REGION Network 15 (SCL): Calculate alarm statuses
   #ST_xStoppingFaults :=  #tALM.tS.xAxisNotAvail OR 
                               #tALM.tS.xInpInstallation OR 
                               #tALM.tS.xAuxPower OR 
                               #tALM.tS.xAreaSafety OR 
                               #tALM.tS.xOverstroke OR 
                               #tALM.tS.xExternInputPower OR 
                               #tALM.tS.xCarriageCutOut OR 
                               #tALM.tS.xDriveTrip OR 
                               #tALM.tS.xDriveNotEnabled OR 
                               #tALM.tS.xAxisNotReady OR 
                               #tALM.tS.xDriveNotReady OR 
                               #tALM.tS.xAxisNotSyncro OR 
                               #tALM.tS.xSpare_12 OR 
                               #tALM.tS.xSpare_13 OR 
                               #tALM.tS.xSpare_14 OR 
                               #tALM.tS.xSpare_15 OR 
                               #tALM.tS.xSpare_16 OR 
                               #tALM.tS.xSpare_17 OR 
                               #tALM.tS.xSpare_18 OR 
                               #tALM.tS.xSpare_19 OR 
                               #tALM.tS.xSpare_20 OR 
                               #tALM.tS.xSpare_21 OR 
                               #tALM.tS.xSpare_22 OR 
                               #tALM.tS.xSpare_23 OR 
                               #tALM.tS.xSpare_24 OR 
                               #tALM.tS.xSpare_25 OR 
                               #tALM.tS.xSpare_26 OR 
                               #tALM.tS.xSpare_27 OR 
                               #tALM.tS.xSpare_28 OR 
                               #tALM.tS.xSpare_29 OR 
                               #tALM.tS.xSpare_30 OR 
                               #tALM.tS.xSpare_31;

   #ST_xFaults := #tALM.tF.xSpare_0 OR
   #tALM.tF.xSpare_1 OR
   #tALM.tF.xSpare_2 OR
   #tALM.tF.xSpare_3 OR
   #tALM.tF.xSpare_4 OR
   #tALM.tF.xSpare_5 OR
   #tALM.tF.xSpare_6 OR
   #tALM.tF.xSpare_7 OR
   #tALM.tF.xSpare_8 OR
   #tALM.tF.xSpare_9 OR
   #tALM.tF.xSpare_10 OR
   #tALM.tF.xSpare_11 OR
   #tALM.tS.xSpare_12 OR
   #tALM.tS.xSpare_13 OR
   #tALM.tS.xSpare_14 OR
   #tALM.tS.xSpare_15 OR
   #tALM.tS.xSpare_16 OR
   #tALM.tS.xSpare_17 OR
   #tALM.tS.xSpare_18 OR
   #tALM.tS.xSpare_19 OR
   #tALM.tS.xSpare_20 OR
   #tALM.tS.xSpare_21 OR
   #tALM.tS.xSpare_22 OR
   #tALM.tS.xSpare_23 OR
   #tALM.tS.xSpare_24 OR
   #tALM.tS.xSpare_25 OR
   #tALM.tS.xSpare_26 OR
   #tALM.tS.xSpare_27 OR
   #tALM.tS.xSpare_28 OR
   #tALM.tS.xSpare_29 OR
   #tALM.tS.xSpare_30 OR
   #tALM.tS.xSpare_31;

   #ST_xWarnings := #tALM.tW.xSpare_0 OR
   #tALM.tW.xSpare_1 OR
   #tALM.tW.xSpare_2 OR
   #tALM.tW.xSpare_3 OR
   #tALM.tW.xSpare_4 OR
   #tALM.tW.xSpare_5 OR
   #tALM.tW.xSpare_6 OR
   #tALM.tW.xSpare_7 OR
   #tALM.tW.xSpare_8 OR
   #tALM.tW.xSpare_9 OR
   #tALM.tW.xSpare_10 OR
   #tALM.tW.xSpare_11 OR
   #tALM.tW.xSpare_12 OR
   #tALM.tW.xSpare_13 OR
   #tALM.tW.xSpare_14 OR
   #tALM.tW.xSpare_15 OR
   #tALM.tW.xSpare_16 OR
   #tALM.tW.xSpare_17 OR
   #tALM.tW.xSpare_18 OR
   #tALM.tW.xSpare_19 OR
   #tALM.tW.xSpare_20 OR
   #tALM.tW.xSpare_21 OR
   #tALM.tW.xSpare_22 OR
   #tALM.tW.xSpare_23 OR
   #tALM.tW.xSpare_24 OR
   #tALM.tW.xSpare_25 OR
   #tALM.tW.xSpare_26 OR
   #tALM.tW.xSpare_27 OR
   #tALM.tW.xSpare_28 OR
   #tALM.tW.xSpare_29 OR
   #tALM.tW.xSpare_30 OR
   #tALM.tW.xSpare_31;
END_REGION

REGION Network 16: Output enable
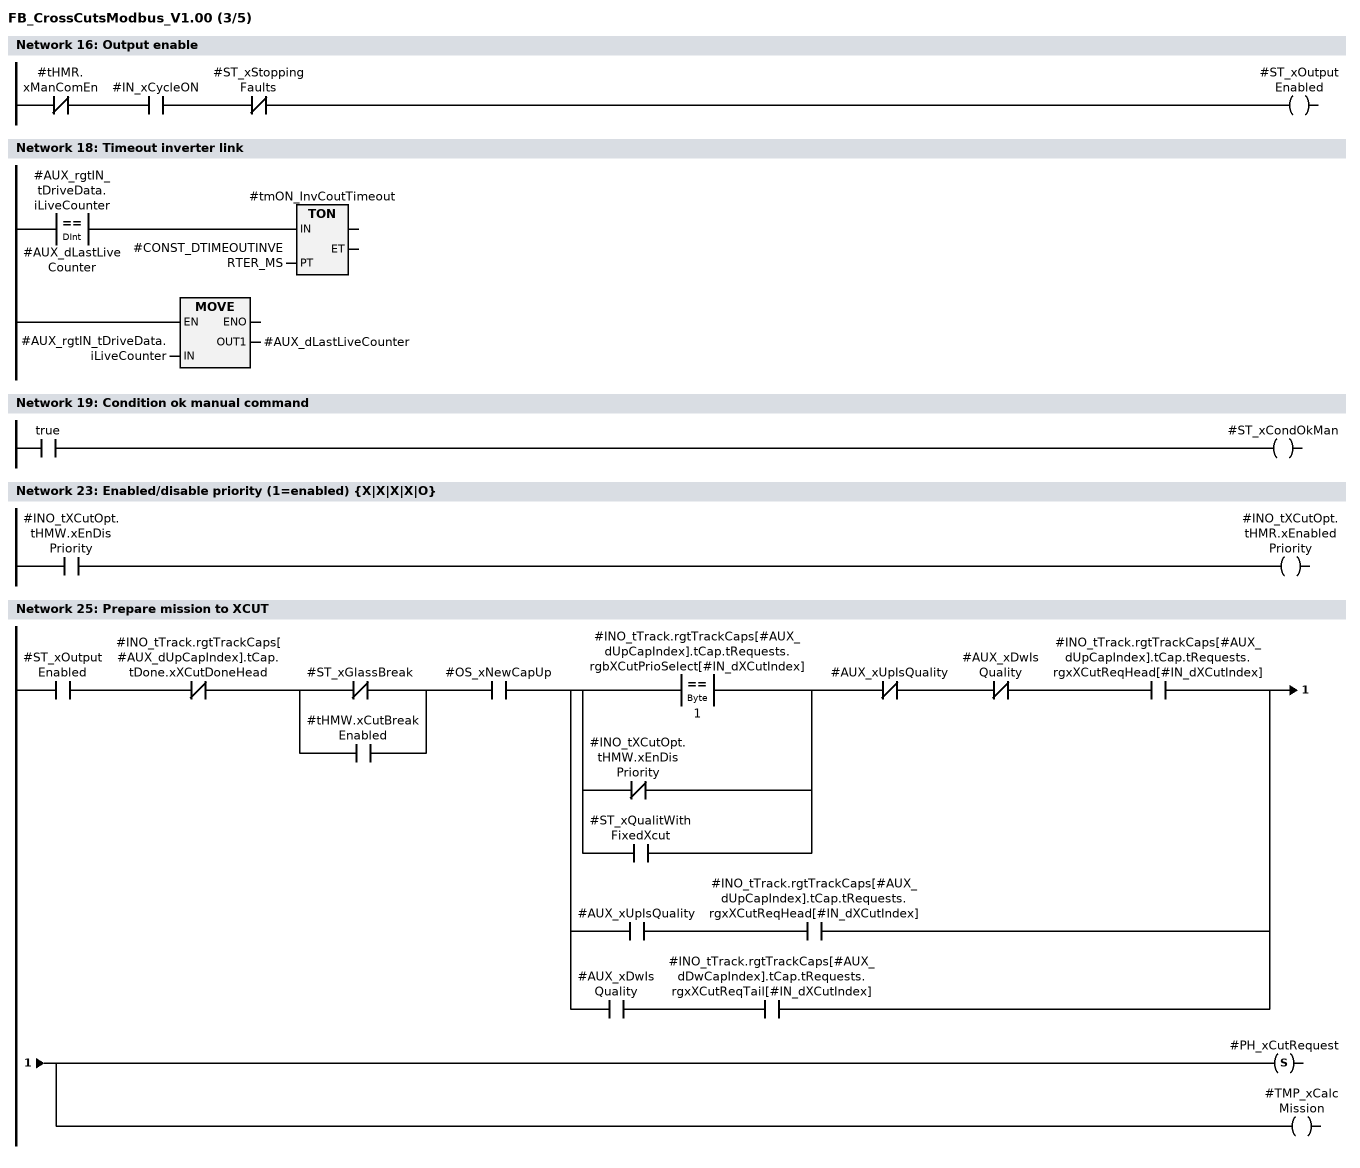
   RUNG wire#powerrail
      I_Contact( #tHMR.xManComEn )
      Contact( #IN_xCycleON )
      I_Contact( #ST_xStoppingFaults )
      Coil( #ST_xOutputEnabled )
   END_RUNG
   // the same network as SCL:
   #ST_xOutputEnabled := NOT #tHMR.xManComEn AND #IN_xCycleON AND NOT #ST_xStoppingFaults;
END_REGION

REGION Network 17 (SCL): Glass break calculation
   #INO_tRibbon.rgtGlassBreakRequest[#IN_dGlassBreakMachineIndex].IN_dDistanceSnaproll_cmm := #tHMR.dDistanceFromSnaproll_cmm;
   #INO_tRibbon.rgtGlassBreakRequest[#IN_dGlassBreakMachineIndex].IN_dDownstreamOffset_cmm := #CONST_DBREAKDOWNOFF_CMM;
   #INO_tRibbon.rgtGlassBreakRequest[#IN_dGlassBreakMachineIndex].IN_dUpstreamOffset_cmm := #CONST_DBREAKUPOFF_CMM;

   IF #INO_tRibbon.rgtGlassBreakRequest[#IN_dGlassBreakMachineIndex].OUT_xDataReady THEN
       #ST_xGlassBreak := #INO_tRibbon.rgtGlassBreakRequest[#IN_dGlassBreakMachineIndex].OUT_xGlassBreak;
   END_IF;

   IF #INO_tRibbon.rgtGlassBreakRequest[#IN_dGlassBreakMachineIndex].OUT_xDataReady OR NOT #INO_tRibbon.rgtGlassBreakRequest[#IN_dGlassBreakMachineIndex].IN_xRequestGlassBreak THEN
       #INO_tRibbon.rgtGlassBreakRequest[#IN_dGlassBreakMachineIndex].OUT_xDataReady := FALSE;
       #INO_tRibbon.rgtGlassBreakRequest[#IN_dGlassBreakMachineIndex].IN_xRequestGlassBreak := TRUE;
   END_IF;
END_REGION

REGION Network 18: Timeout inverter link
   #tmON_InvCoutTimeout(IN := #AUX_rgtIN_tDriveData.iLiveCounter = #AUX_dLastLiveCounter,   // TON
                        PT := #CONST_DTIMEOUTINVERTER_MS);
   #AUX_dLastLiveCounter := #AUX_rgtIN_tDriveData.iLiveCounter;
END_REGION

REGION Network 19: Condition ok manual command
   RUNG wire#powerrail
      Contact( true )
      Coil( #ST_xCondOkMan )
   END_RUNG
   // the same network as SCL:
   #ST_xCondOkMan := true;
END_REGION

REGION Network 20: ####_PHASES_&_LOGICS_####
END_REGION

REGION Network 21 (SCL): Calculate return speed
   IF #PH_xEndCutRequest AND #AUX_xValidUpCap THEN
       #TMP_dCutYSpace_cmm := #AUX_dCutStopPosUp_cmm;

       #TMP_dCutSpace_cmm := REAL_TO_DINT(DINT_TO_REAL(#TMP_dCutYSpace_cmm) * (TAN(((3.14 * (DINT_TO_REAL(#tHMR.dAngleValue_uDegree) / 1000000.0)) / 180.0))));

       #AUX_dSimStoreCutTime_ms := #TMP_dCutTime_ms := REAL_TO_DINT((DINT_TO_REAL(#TMP_dCutSpace_cmm + 30000)) / #INO_tEnc.rActSpeedValue_cmm_ms);

       #AUX_dSimCutSpace_cmm := #TMP_dTravSpace_cmm :=  REAL_TO_DINT(SQRT(((DINT_TO_REAL(#TMP_dCutYSpace_cmm) / 100) ** 2) + ((DINT_TO_REAL(#TMP_dCutSpace_cmm) / 100) ** 2))) * 100 + 36000;

       //Calculate at 20%

       #TMP_rAccTime_s := ((DINT_TO_REAL(#CONST_DSPEED_CMM_S) * 0.2)) / DINT_TO_REAL(#CONST_DRAMP_CMM_S2);

       #TMP_dRampSpace_cmm := REAL_TO_DINT((((#TMP_rAccTime_s ** 2) * 0.5) * DINT_TO_REAL(#CONST_DRAMP_CMM_S2)) * 2);

       #TMP_dConstSpace_cmm := #TMP_dTravSpace_cmm - #TMP_dRampSpace_cmm;
       #TMP_dConstTime_ms := REAL_TO_DINT(((DINT_TO_REAL(#TMP_dConstSpace_cmm) / (DINT_TO_REAL(#CONST_DSPEED_CMM_S) * 0.2))) * 1000.0);

       #AUX_dCutTime20Per_ms := #TMP_dCutTime_ms + #TMP_dConstTime_ms + REAL_TO_DINT(((#TMP_rAccTime_s * 1000) * 2));

       //Calculate at 40%

       #TMP_rAccTime_s := ((DINT_TO_REAL(#CONST_DSPEED_CMM_S) * 0.4)) / DINT_TO_REAL(#CONST_DRAMP_CMM_S2);

       #TMP_dRampSpace_cmm := REAL_TO_DINT((((#TMP_rAccTime_s ** 2) * 0.5) * DINT_TO_REAL(#CONST_DRAMP_CMM_S2)) * 2);

       #TMP_dConstSpace_cmm := #TMP_dTravSpace_cmm - #TMP_dRampSpace_cmm;
       #TMP_dConstTime_ms := REAL_TO_DINT(((DINT_TO_REAL(#TMP_dConstSpace_cmm) / (DINT_TO_REAL(#CONST_DSPEED_CMM_S) * 0.4))) * 1000.0);

       #AUX_dCutTime40Per_ms := #TMP_dCutTime_ms + #TMP_dConstTime_ms + REAL_TO_DINT(((#TMP_rAccTime_s * 1000) * 2));

       //Calculate at 60%

       #TMP_rAccTime_s := ((DINT_TO_REAL(#CONST_DSPEED_CMM_S) * 0.6)) / DINT_TO_REAL(#CONST_DRAMP_CMM_S2);

       #TMP_dRampSpace_cmm := REAL_TO_DINT((((#TMP_rAccTime_s ** 2) * 0.5) * DINT_TO_REAL(#CONST_DRAMP_CMM_S2)) * 2);

       #TMP_dConstSpace_cmm := #TMP_dTravSpace_cmm - #TMP_dRampSpace_cmm;
       #TMP_dConstTime_ms := (REAL_TO_DINT(((DINT_TO_REAL(#TMP_dConstSpace_cmm) / (DINT_TO_REAL(#CONST_DSPEED_CMM_S) * 0.6))) * 1000.0));

       #AUX_dCutTime60Per_ms := #TMP_dCutTime_ms + #TMP_dConstTime_ms + REAL_TO_DINT(((#TMP_rAccTime_s * 1000) * 2));

       //Calculate at 80%

       #TMP_rAccTime_s := ((DINT_TO_REAL(#CONST_DSPEED_CMM_S) * 0.8)) / DINT_TO_REAL(#CONST_DRAMP_CMM_S2);

       #TMP_dRampSpace_cmm := REAL_TO_DINT((((#TMP_rAccTime_s ** 2) * 0.5) * DINT_TO_REAL(#CONST_DRAMP_CMM_S2)) * 2);

       #TMP_dConstSpace_cmm := #TMP_dTravSpace_cmm - #TMP_dRampSpace_cmm;
       #TMP_dConstTime_ms := REAL_TO_DINT(((DINT_TO_REAL(#TMP_dConstSpace_cmm) / (DINT_TO_REAL(#CONST_DSPEED_CMM_S) * 0.8))) * 1000.0);

       #AUX_dCutTime80Per_ms := #TMP_dCutTime_ms + #TMP_dConstTime_ms + REAL_TO_DINT(((#TMP_rAccTime_s * 1000) * 2));

       //Calculate at 100%
       #TMP_rAccTime_s := ((DINT_TO_REAL(#CONST_DSPEED_CMM_S) * 1.0)) / DINT_TO_REAL(#CONST_DRAMP_CMM_S2);

       #TMP_dRampSpace_cmm := REAL_TO_DINT((((#TMP_rAccTime_s ** 2) * 0.5) * DINT_TO_REAL(#CONST_DRAMP_CMM_S2)) * 2);

       #TMP_dConstSpace_cmm := #TMP_dTravSpace_cmm - #TMP_dRampSpace_cmm;
       #TMP_dConstTime_ms := REAL_TO_DINT(((DINT_TO_REAL(#TMP_dConstSpace_cmm) / (DINT_TO_REAL(#CONST_DSPEED_CMM_S) * 1.0))) * 1000.0);
       #AUX_dCutTime100Per_ms := #TMP_dCutTime_ms + #TMP_dConstTime_ms + REAL_TO_DINT(((#TMP_rAccTime_s * 1000) * 2));


       //Calculate next plate time
       #AUX_dNextPlateTime_ms := REAL_TO_DINT((DINT_TO_REAL(#INO_tTrack.rgtTrackCaps[#AUX_dUpCapIndex].tCap.dLength_cmm - 50000)) / #INO_tEnc.rActSpeedValue_cmm_ms);
   END_IF;
END_REGION

REGION Network 22 (SCL): Calculate positions

   IF #OS_xNewCap THEN

       #AUX_dCutStartPosUp_cmm := #CONST_DMAXCUTRANGE_CMM;
       #AUX_dCutStartPosDw_cmm := #CONST_DMAXCUTRANGE_CMM;

       #AUX_dCutStopPosUp_cmm := #CONST_DMINCUTRANGE_CMM;
       #AUX_dCutStopPosDw_cmm := #CONST_DMINCUTRANGE_CMM;

       CASE #tHMR.dActualCutPosRequest OF

           #CONST_DMODECUT_OPERATOR:
               #AUX_dCutStartPosUp_cmm :=ABS_DINT(#tHMR.dDistanceFromCenterLine_cmm) + #tHMW.dOperStartCutPos_cmm + #tHMW.dCutStartOffsetDelay_cmm;
               #AUX_dCutStopPosUp_cmm := ABS_DINT(#tHMR.dDistanceFromCenterLine_cmm) + #tHMW.dOperEndCutPos_cmm + #tHMW.dCutEndOffsetDelay_cmm;

               #AUX_dCutStartPosDw_cmm := ABS_DINT(#tHMR.dDistanceFromCenterLine_cmm) +#tHMW.dOperStartCutPos_cmm + #tHMW.dCutStartOffsetDelay_cmm;
               #AUX_dCutStopPosDw_cmm := ABS_DINT(#tHMR.dDistanceFromCenterLine_cmm) + #tHMW.dOperEndCutPos_cmm + #tHMW.dCutEndOffsetDelay_cmm;

           #CONST_DMODECUT_GROSS:
               IF #OS_xNewCapUp THEN
                   #AUX_dCutStartPosUp_cmm := ABS_DINT(#tHMR.dDistanceFromCenterLine_cmm) + (#INO_tTrack.rgtTrackCaps[#AUX_dUpCapIndex].tCap.dGrossWidth_cmm / -2) +
                                                #INO_tTrack.rgtTrackCaps[#AUX_dUpCapIndex].tCap.dGrossWander_cmm +  #tHMW.dCutStartOffsetDelay_cmm;
                   #AUX_dCutStopPosUp_cmm := ABS_DINT(#tHMR.dDistanceFromCenterLine_cmm) + (#INO_tTrack.rgtTrackCaps[#AUX_dUpCapIndex].tCap.dGrossWidth_cmm / 2) +
                                                #INO_tTrack.rgtTrackCaps[#AUX_dUpCapIndex].tCap.dGrossWander_cmm +  #tHMW.dCutEndOffsetDelay_cmm;
               END_IF;

               IF #OS_xNewCapDw THEN
                   #AUX_dCutStartPosDw_cmm := ABS_DINT(#tHMR.dDistanceFromCenterLine_cmm) + (#INO_tTrack.rgtTrackCaps[#AUX_dDwCapIndex].tCap.dGrossWidth_cmm / -2) +
                                                #INO_tTrack.rgtTrackCaps[#AUX_dDwCapIndex].tCap.dGrossWander_cmm +  #tHMW.dCutStartOffsetDelay_cmm;
                   #AUX_dCutStopPosDw_cmm := ABS_DINT(#tHMR.dDistanceFromCenterLine_cmm) + (#INO_tTrack.rgtTrackCaps[#AUX_dDwCapIndex].tCap.dGrossWidth_cmm / 2) +
                                                #INO_tTrack.rgtTrackCaps[#AUX_dDwCapIndex].tCap.dGrossWander_cmm +  #tHMW.dCutEndOffsetDelay_cmm;
               END_IF;

           #CONST_DMODECUT_NET:
               IF #OS_xNewCapUp THEN
                   #AUX_dCutStartPosUp_cmm := ABS_DINT(#tHMR.dDistanceFromCenterLine_cmm) + (#INO_tTrack.rgtTrackCaps[#AUX_dUpCapIndex].tCap.dNetWidth_cmm / -2) +
                                                #INO_tTrack.rgtTrackCaps[#AUX_dUpCapIndex].tCap.dNetWander_cmm +  #tHMW.dCutStartOffsetDelay_cmm;
                   #AUX_dCutStopPosUp_cmm := ABS_DINT(#tHMR.dDistanceFromCenterLine_cmm) + (#INO_tTrack.rgtTrackCaps[#AUX_dUpCapIndex].tCap.dNetWidth_cmm / 2) +
                                                    #INO_tTrack.rgtTrackCaps[#AUX_dUpCapIndex].tCap.dNetWander_cmm +  #tHMW.dCutEndOffsetDelay_cmm;
               END_IF;

               IF #OS_xNewCapDw THEN
                   #AUX_dCutStartPosDw_cmm := ABS_DINT(#tHMR.dDistanceFromCenterLine_cmm) + (#INO_tTrack.rgtTrackCaps[#AUX_dDwCapIndex].tCap.dNetWidth_cmm / -2) +
                                                #INO_tTrack.rgtTrackCaps[#AUX_dDwCapIndex].tCap.dNetWander_cmm +  #tHMW.dCutStartOffsetDelay_cmm;
                   #AUX_dCutStopPosDw_cmm := ABS_DINT(#tHMR.dDistanceFromCenterLine_cmm) + (#INO_tTrack.rgtTrackCaps[#AUX_dDwCapIndex].tCap.dNetWidth_cmm / 2) +
                                                    #INO_tTrack.rgtTrackCaps[#AUX_dDwCapIndex].tCap.dNetWander_cmm +  #tHMW.dCutEndOffsetDelay_cmm;
               END_IF;

           #CONST_DMODECUT_YCUT:
               IF #OS_xNewCapUp THEN
                   #AUX_dCutStartPosUp_cmm := ABS_DINT(#tHMR.dDistanceFromCenterLine_cmm) + (#INO_tTrack.rgtTrackCaps[#AUX_dUpCapIndex].tCap.dWidth_cmm / -2) +
                                                #INO_tTrack.rgtTrackCaps[#AUX_dUpCapIndex].tCap.dStartCutWander_cmm +  #tHMW.dCutStartOffsetDelay_cmm;
                   #AUX_dCutStopPosUp_cmm := ABS_DINT(#tHMR.dDistanceFromCenterLine_cmm) + (#INO_tTrack.rgtTrackCaps[#AUX_dUpCapIndex].tCap.dWidth_cmm / 2) +
                                                #INO_tTrack.rgtTrackCaps[#AUX_dUpCapIndex].tCap.dStartCutWander_cmm +  #tHMW.dCutEndOffsetDelay_cmm;
               END_IF;

               IF #OS_xNewCapDw THEN
                   #AUX_dCutStartPosDw_cmm := ABS_DINT(#tHMR.dDistanceFromCenterLine_cmm) + (#INO_tTrack.rgtTrackCaps[#AUX_dDwCapIndex].tCap.dWidth_cmm / -2) +
                                                #INO_tTrack.rgtTrackCaps[#AUX_dDwCapIndex].tCap.dStartCutWander_cmm +  #tHMW.dCutStartOffsetDelay_cmm;
                   #AUX_dCutStopPosDw_cmm := ABS_DINT(#tHMR.dDistanceFromCenterLine_cmm) + (#INO_tTrack.rgtTrackCaps[#AUX_dDwCapIndex].tCap.dWidth_cmm / 2) +
                                                #INO_tTrack.rgtTrackCaps[#AUX_dDwCapIndex].tCap.dStartCutWander_cmm +  #tHMW.dCutEndOffsetDelay_cmm;
               END_IF;


       END_CASE;


   END_IF;
END_REGION

REGION Network 23: Enabled/disable priority (1=enabled) {X|X|X|X|O}
   RUNG wire#powerrail
      Contact( #INO_tXCutOpt.tHMW.xEnDisPriority )
      Coil( #INO_tXCutOpt.tHMR.xEnabledPriority )
   END_RUNG
   // the same network as SCL:
   #INO_tXCutOpt.tHMR.xEnabledPriority := #INO_tXCutOpt.tHMW.xEnDisPriority;
END_REGION

REGION Network 24 (SCL): Priority manager

   #INO_tXCutOpt.IN_rgdCutTime_ms[#IN_dXCutIndex] := #AUX_dCutTime100Per_ms;
   #INO_tXCutOpt.IN_rgxCutsAvailable[#IN_dXCutIndex] := (#tHMR.dXCutActualStatus=3);
   #INO_tXCutOpt.IN_rgdPiorityList[#IN_dXCutIndex] := #tHMW.dCutPriority;
   #INO_tXCutOpt(IN_dActualNumOfXCuts :="DMAXXHEADS",
                                   IN_dCapIndexCall := #AUX_dUpCapIndex,
                                   IN_dXCutCallIndex := #IN_dXCutIndex,
                                   IN_xNewTargetCall := #OS_xNewCap,
                                   IN_xRescueCall := false,
                                   INO_tOBInit := "GP_OB_Initialize_Slow_IDB",
                                   INO_tTrack:=#INO_tTrack);

   IF #OS_xNewCap THEN
                         #ST_xQualitWithFixedXcut := 0;
                         #INO_tTrack.rgtTrackSearch[#IN_dGlassSearchMachineIndex_Q0].xPlateFound := 0;
                         #INO_tTrack.rgtTrackSearch[#IN_dGlassSearchMachineIndex_Q0].xRequestSearchPlate := 1;
                         #INO_tTrack.rgtTrackSearch[#IN_dGlassSearchMachineIndex_Q0].dSearchMode := 2;
                         #INO_tTrack.rgtTrackSearch[#IN_dGlassSearchMachineIndex_Q0].dRequestID += 1;
                         #INO_tTrack.rgtTrackSearch[#IN_dGlassSearchMachineIndex_Q0].dMaxTailPosition_cmm := #tHMR.dDistanceFromSnaproll_cmm + 1000000;
                         #INO_tTrack.rgtTrackSearch[#IN_dGlassSearchMachineIndex_Q0].dMinTailPosition_cmm := #tHMR.dDistanceFromSnaproll_cmm - 400000;
                         #INO_tTrack.rgtTrackSearch[#IN_dGlassSearchMachineIndex_Q0].tSearchRequest.xMainDestEqual := 1;
                         #INO_tTrack.rgtTrackSearch[#IN_dGlassSearchMachineIndex_Q0].tSearchData.dMainDest_mask := "DQUALITYDESTMASK1";

                         #INO_tTrack.rgtTrackSearch[#IN_dGlassSearchMachineIndex_Q1].xPlateFound := 0;
                         #INO_tTrack.rgtTrackSearch[#IN_dGlassSearchMachineIndex_Q1].xRequestSearchPlate := 1;
                         #INO_tTrack.rgtTrackSearch[#IN_dGlassSearchMachineIndex_Q1].dSearchMode := 2;
                         #INO_tTrack.rgtTrackSearch[#IN_dGlassSearchMachineIndex_Q1].dRequestID += 1;
                         #INO_tTrack.rgtTrackSearch[#IN_dGlassSearchMachineIndex_Q1].dMaxTailPosition_cmm := #tHMR.dDistanceFromSnaproll_cmm + 1000000;
                         #INO_tTrack.rgtTrackSearch[#IN_dGlassSearchMachineIndex_Q1].dMinTailPosition_cmm := #tHMR.dDistanceFromSnaproll_cmm - 400000;
                         #INO_tTrack.rgtTrackSearch[#IN_dGlassSearchMachineIndex_Q1].tSearchRequest.xMainDestEqual := 1;
                         #INO_tTrack.rgtTrackSearch[#IN_dGlassSearchMachineIndex_Q1].tSearchData.dMainDest_mask := "DQUALITYDESTMASK2";

                         #INO_tTrack.rgtTrackSearch[#IN_dGlassSearchMachineIndex_Q2].xPlateFound := 0;
                         #INO_tTrack.rgtTrackSearch[#IN_dGlassSearchMachineIndex_Q2].xRequestSearchPlate := 1;
                         #INO_tTrack.rgtTrackSearch[#IN_dGlassSearchMachineIndex_Q2].dSearchMode := 2;
                         #INO_tTrack.rgtTrackSearch[#IN_dGlassSearchMachineIndex_Q2].dRequestID += 1;
                         #INO_tTrack.rgtTrackSearch[#IN_dGlassSearchMachineIndex_Q2].dMaxTailPosition_cmm := #tHMR.dDistanceFromSnaproll_cmm + 1000000;
                         #INO_tTrack.rgtTrackSearch[#IN_dGlassSearchMachineIndex_Q2].dMinTailPosition_cmm := #tHMR.dDistanceFromSnaproll_cmm - 400000;
                         #INO_tTrack.rgtTrackSearch[#IN_dGlassSearchMachineIndex_Q2].tSearchRequest.xMainDestEqual := 1;
                         #INO_tTrack.rgtTrackSearch[#IN_dGlassSearchMachineIndex_Q2].tSearchData.dMainDest_mask := "DQUALITYDESTMASK3";

                         #INO_tTrack.rgtTrackSearch[#IN_dGlassSearchMachineIndex_Q2].xPlateFound := 0;
                         #INO_tTrack.rgtTrackSearch[#IN_dGlassSearchMachineIndex_Q2].xRequestSearchPlate := 1;
                         #INO_tTrack.rgtTrackSearch[#IN_dGlassSearchMachineIndex_Q2].dSearchMode := 2;
                         #INO_tTrack.rgtTrackSearch[#IN_dGlassSearchMachineIndex_Q2].dRequestID += 1;
                         #INO_tTrack.rgtTrackSearch[#IN_dGlassSearchMachineIndex_Q2].dMaxTailPosition_cmm := #tHMR.dDistanceFromSnaproll_cmm + 1000000;
                         #INO_tTrack.rgtTrackSearch[#IN_dGlassSearchMachineIndex_Q2].dMinTailPosition_cmm := #tHMR.dDistanceFromSnaproll_cmm - 400000;
                         #INO_tTrack.rgtTrackSearch[#IN_dGlassSearchMachineIndex_Q2].tSearchRequest.xMainDestEqual := 1;
                         #INO_tTrack.rgtTrackSearch[#IN_dGlassSearchMachineIndex_Q2].tSearchData.dMainDest_mask := "DQUALITYDESTMASK4";
   END_IF;

   IF #INO_tTrack.rgtTrackSearch[#IN_dGlassSearchMachineIndex_Q0].xPlateFound OR #INO_tTrack.rgtTrackSearch[#IN_dGlassSearchMachineIndex_Q1].xPlateFound OR #INO_tTrack.rgtTrackSearch[#IN_dGlassSearchMachineIndex_Q2].xPlateFound THEN
       FOR #TMP_dIndex := 0 TO "DMAXXHEADS" - 1 DO
           IF #INO_tTrack.rgtTrackCaps[#INO_tTrack.rgtTrackSearch[#IN_dGlassSearchMachineIndex_Q0].dFoundTrackIndex].tCap.tRequests.rgxXCutReqHead[#TMP_dIndex] = 0 THEN
               #ST_xQualitWithFixedXcut := 1;
           END_IF;
       END_FOR;
   END_IF;
END_REGION

REGION Network 25: Prepare mission to XCUT
   RUNG wire#powerrail
      Contact( #ST_xOutputEnabled )
      I_Contact( #INO_tTrack.rgtTrackCaps[#AUX_dUpCapIndex].tCap.tDone.xXCutDoneHead )
      wire#w1
      I_Contact( #ST_xGlassBreak )
      wire#w2
      Contact( #OS_xNewCapUp )
      wire#w3
      { S7_Templates := "SrcType := Byte" } EQ_Contact(in1 := #INO_tTrack.rgtTrackCaps[#AUX_dUpCapIndex].tCap.tRequests.rgbXCutPrioSelect[#IN_dXCutIndex], in2 := 1)
      wire#w4
      I_Contact( #AUX_xUpIsQuality )
      I_Contact( #AUX_xDwIsQuality )
      Contact( #INO_tTrack.rgtTrackCaps[#AUX_dUpCapIndex].tCap.tRequests.rgxXCutReqHead[#IN_dXCutIndex] )
      wire#w5
      S_Coil( #PH_xCutRequest )
   END_RUNG
   RUNG wire#w1
      Contact( #tHMW.xCutBreakEnabled )
   END_RUNG wire#w2
   RUNG wire#w3
      I_Contact( #INO_tXCutOpt.tHMW.xEnDisPriority )
   END_RUNG wire#w4
   RUNG wire#w3
      Contact( #ST_xQualitWithFixedXcut )
   END_RUNG wire#w4
   RUNG wire#w3
      Contact( #AUX_xUpIsQuality )
      Contact( #INO_tTrack.rgtTrackCaps[#AUX_dUpCapIndex].tCap.tRequests.rgxXCutReqHead[#IN_dXCutIndex] )
   END_RUNG wire#w5
   RUNG wire#w3
      Contact( #AUX_xDwIsQuality )
      Contact( #INO_tTrack.rgtTrackCaps[#AUX_dDwCapIndex].tCap.tRequests.rgxXCutReqTail[#IN_dXCutIndex] )
   END_RUNG wire#w5
   RUNG wire#w5
      Coil( #TMP_xCalcMission )
   END_RUNG
   // the same network as SCL:
   #_w1 := #ST_xOutputEnabled AND NOT #INO_tTrack.rgtTrackCaps[#AUX_dUpCapIndex].tCap.tDone.xXCutDoneHead AND (NOT #ST_xGlassBreak OR #tHMW.xCutBreakEnabled) AND #OS_xNewCapUp AND ((((#INO_tTrack.rgtTrackCaps[#AUX_dUpCapIndex].tCap.tRequests.rgbXCutPrioSelect[#IN_dXCutIndex] = 1) OR NOT #INO_tXCutOpt.tHMW.xEnDisPriority OR #ST_xQualitWithFixedXcut) AND NOT #AUX_xUpIsQuality AND NOT #AUX_xDwIsQuality AND #INO_tTrack.rgtTrackCaps[#AUX_dUpCapIndex].tCap.tRequests.rgxXCutReqHead[#IN_dXCutIndex]) OR (#AUX_xUpIsQuality AND #INO_tTrack.rgtTrackCaps[#AUX_dUpCapIndex].tCap.tRequests.rgxXCutReqHead[#IN_dXCutIndex]) OR (#AUX_xDwIsQuality AND #INO_tTrack.rgtTrackCaps[#AUX_dDwCapIndex].tCap.tRequests.rgxXCutReqTail[#IN_dXCutIndex]));
   IF #_w1 THEN #PH_xCutRequest := TRUE; END_IF;
   #TMP_xCalcMission := #_w1;
END_REGION

REGION Network 26 (SCL): Prepare data for the new mission
   IF #TMP_xCalcMission THEN

       #AUX_dMissionToSend := #AUX_dMissionToSend + 1;

       IF #AUX_dMissionToSend > #CONST_DMAXMISSIONNUM THEN
           #AUX_dMissionToSend := 1;
       END_IF;

       #AUX_dMissionCounterValue_cmm := #INO_tTrack.rgtTrackMachine[#IN_dMachineIndex].tUserData.dGetEncValueOnSnap_cmm - #tHMR.dDistanceFromSnaproll_cmm + #tHMW.dPosOffset_cmm;

       IF (#IN_xSimulationActive) THEN

           #AUX_rgtIN_tDriveData.dMissionDone := 0;

           IF (#AUX_dSimWaitEnd_ms <= 0) THEN
               //The bridge is free can assign this cut
               #AUX_rgtIN_tDriveData.dMissionDone := #AUX_dMissionToSend;
               #AUX_dSimWaitEnd_ms := #AUX_dCutTime100Per_ms;
               #AUX_dSimCutTime_ms := #AUX_dSimStoreCutTime_ms;
           ELSE
               #AUX_rgtIN_tDriveData.dMissionUnDone := #AUX_dMissionToSend;
           END_IF;        
       END_IF;
   END_IF;
END_REGION

REGION Network 27 (SCL): Decrease simulation incutting counter
   IF (#IN_xSimulationActive) THEN

       #AUX_dSimWaitEnd_ms -= #INO_tOBInit.OUT_dExecutionTime_ms;
       #AUX_dSimCutTime_ms -= #INO_tOBInit.OUT_dExecutionTime_ms;

       IF (#AUX_dSimWaitEnd_ms < 0) THEN
           #AUX_dSimWaitEnd_ms := 0;
       END_IF;

       IF (#AUX_dSimCutTime_ms < 0) THEN
           #AUX_dSimCutTime_ms := 0;
       END_IF;

       //Calculate the carriage position in according to the cutting time
       IF #AUX_dSimCutTime_ms > 0 THEN
           #tHMR.dCarriagePosition_cmm := REAL_TO_DINT(DINT_TO_REAL(#AUX_dSimCutSpace_cmm) * (DINT_TO_REAL(#AUX_dSimStoreCutTime_ms - #AUX_dSimCutTime_ms) / DINT_TO_REAL(#AUX_dSimStoreCutTime_ms)));
       ELSE
           #tHMR.dCarriagePosition_cmm := REAL_TO_DINT(DINT_TO_REAL(#AUX_dSimCutSpace_cmm) * (DINT_TO_REAL(#AUX_dSimWaitEnd_ms) / DINT_TO_REAL(#AUX_dCutTime100Per_ms - #AUX_dSimStoreCutTime_ms)));

       END_IF;

   END_IF;
END_REGION

REGION Network 28: End cut request
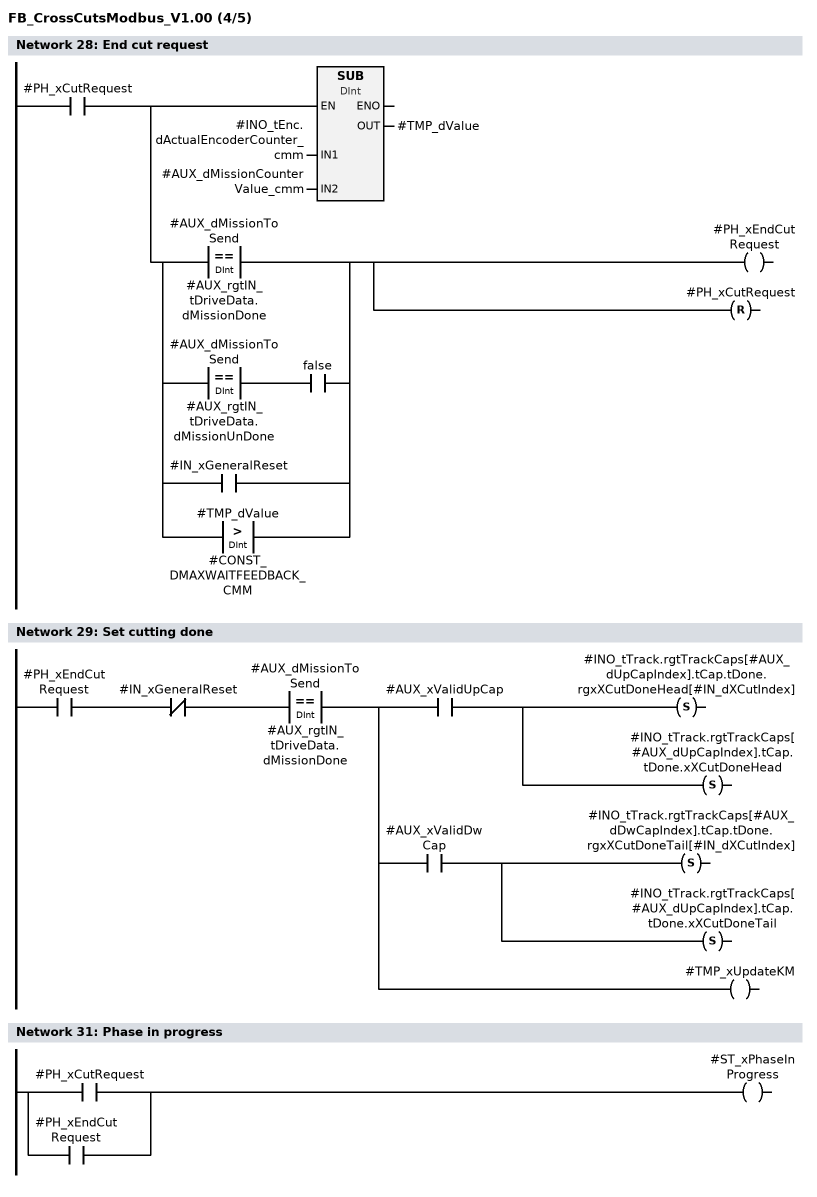
   RUNG wire#powerrail
      Contact( #PH_xCutRequest )
      wire#w1
      { S7_Templates := "SrcType := DInt" } Sub(in1 := #INO_tEnc.dActualEncoderCounter_cmm, in2 := #AUX_dMissionCounterValue_cmm, out => #TMP_dValue)
   END_RUNG
   RUNG wire#w1
      { S7_Templates := "SrcType := DInt" } EQ_Contact(in1 := #AUX_dMissionToSend, in2 := #AUX_rgtIN_tDriveData.dMissionDone)
      wire#w2
      Coil( #PH_xEndCutRequest )
   END_RUNG
   RUNG wire#w1
      { S7_Templates := "SrcType := DInt" } EQ_Contact(in1 := #AUX_dMissionToSend, in2 := #AUX_rgtIN_tDriveData.dMissionUnDone)
      Contact( false )
   END_RUNG wire#w2
   RUNG wire#w1
      Contact( #IN_xGeneralReset )
   END_RUNG wire#w2
   RUNG wire#w1
      { S7_Templates := "SrcType := DInt" } GT_Contact(in1 := #TMP_dValue, in2 := #CONST_DMAXWAITFEEDBACK_CMM)
   END_RUNG wire#w2
   RUNG wire#w2
      R_Coil( #PH_xCutRequest )
   END_RUNG
   // the same network as SCL:
   IF #PH_xCutRequest THEN
       #TMP_dValue := #INO_tEnc.dActualEncoderCounter_cmm - #AUX_dMissionCounterValue_cmm;
   END_IF;
   #PH_xEndCutRequest := #PH_xCutRequest AND ((#AUX_dMissionToSend = #AUX_rgtIN_tDriveData.dMissionDone) OR ((#AUX_dMissionToSend = #AUX_rgtIN_tDriveData.dMissionUnDone) AND false) OR #IN_xGeneralReset OR (#TMP_dValue > #CONST_DMAXWAITFEEDBACK_CMM));
   IF #PH_xEndCutRequest THEN #PH_xCutRequest := FALSE; END_IF;
END_REGION

REGION Network 29: Set cutting done
   RUNG wire#powerrail
      Contact( #PH_xEndCutRequest )
      I_Contact( #IN_xGeneralReset )
      { S7_Templates := "SrcType := DInt" } EQ_Contact(in1 := #AUX_dMissionToSend, in2 := #AUX_rgtIN_tDriveData.dMissionDone)
      wire#w1
      Contact( #AUX_xValidUpCap )
      wire#w2
      S_Coil( #INO_tTrack.rgtTrackCaps[#AUX_dUpCapIndex].tCap.tDone.rgxXCutDoneHead[#IN_dXCutIndex] )
   END_RUNG
   RUNG wire#w2
      S_Coil( #INO_tTrack.rgtTrackCaps[#AUX_dUpCapIndex].tCap.tDone.xXCutDoneHead )
   END_RUNG
   RUNG wire#w1
      Contact( #AUX_xValidDwCap )
      wire#w3
      S_Coil( #INO_tTrack.rgtTrackCaps[#AUX_dDwCapIndex].tCap.tDone.rgxXCutDoneTail[#IN_dXCutIndex] )
   END_RUNG
   RUNG wire#w3
      S_Coil( #INO_tTrack.rgtTrackCaps[#AUX_dUpCapIndex].tCap.tDone.xXCutDoneTail )
   END_RUNG
   RUNG wire#w1
      Coil( #TMP_xUpdateKM )
   END_RUNG
   // the same network as SCL:
   #_w1 := #PH_xEndCutRequest AND NOT #IN_xGeneralReset AND (#AUX_dMissionToSend = #AUX_rgtIN_tDriveData.dMissionDone);
   IF #_w1 AND #AUX_xValidUpCap THEN
       #INO_tTrack.rgtTrackCaps[#AUX_dUpCapIndex].tCap.tDone.rgxXCutDoneHead[#IN_dXCutIndex] := TRUE;
       #INO_tTrack.rgtTrackCaps[#AUX_dUpCapIndex].tCap.tDone.xXCutDoneHead := TRUE;
   END_IF;
   IF #_w1 AND #AUX_xValidDwCap THEN
       #INO_tTrack.rgtTrackCaps[#AUX_dDwCapIndex].tCap.tDone.rgxXCutDoneTail[#IN_dXCutIndex] := TRUE;
       #INO_tTrack.rgtTrackCaps[#AUX_dUpCapIndex].tCap.tDone.xXCutDoneTail := TRUE;
   END_IF;
   #TMP_xUpdateKM := #_w1;
END_REGION

REGION Network 30 (SCL): Calculate head Km
   IF #TMP_xUpdateKM THEN

       #tHMR.rHeadUsage_km := #tHMR.rHeadUsage_km + DINT_TO_REAL(#tHMW.dOperEndCutPos_cmm - #tHMW.dOperStartCutPos_cmm) / 100000000.0;

   END_IF;
END_REGION

REGION Network 31: Phase in progress
   RUNG wire#powerrail
      Contact( #PH_xCutRequest )
      wire#w1
      Coil( #ST_xPhaseInProgress )
   END_RUNG
   RUNG wire#powerrail
      Contact( #PH_xEndCutRequest )
   END_RUNG wire#w1
   // the same network as SCL:
   #ST_xPhaseInProgress := #PH_xCutRequest OR #PH_xEndCutRequest;
END_REGION

REGION Network 32: Modbus phases
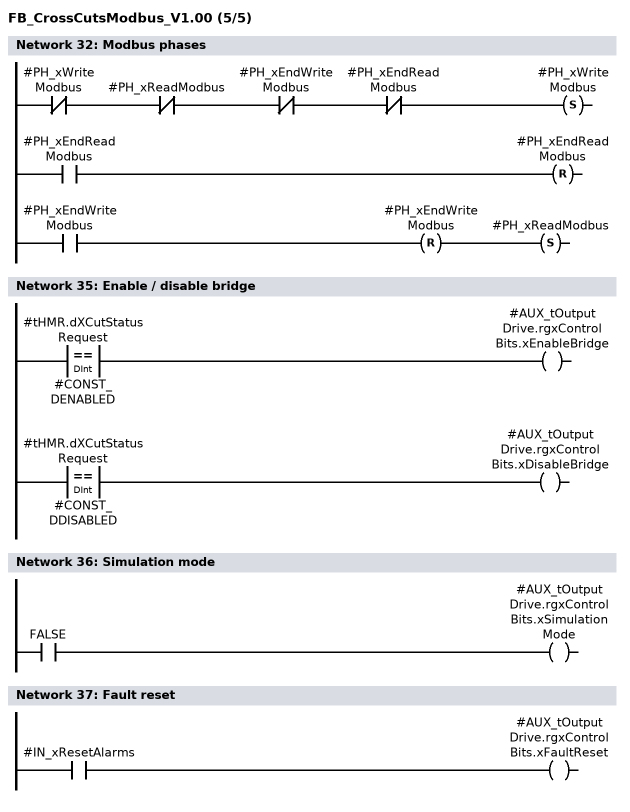
   RUNG wire#powerrail
      I_Contact( #PH_xWriteModbus )
      I_Contact( #PH_xReadModbus )
      I_Contact( #PH_xEndWriteModbus )
      I_Contact( #PH_xEndReadModbus )
      S_Coil( #PH_xWriteModbus )
   END_RUNG
   RUNG wire#powerrail
      Contact( #PH_xEndReadModbus )
      R_Coil( #PH_xEndReadModbus )
   END_RUNG
   RUNG wire#powerrail
      Contact( #PH_xEndWriteModbus )
      R_Coil( #PH_xEndWriteModbus )
      S_Coil( #PH_xReadModbus )
   END_RUNG
   // the same network as SCL:
   IF NOT #PH_xWriteModbus AND NOT #PH_xReadModbus AND NOT #PH_xEndWriteModbus AND NOT #PH_xEndReadModbus THEN
       #PH_xWriteModbus := TRUE;
   END_IF;
   IF #PH_xEndReadModbus THEN #PH_xEndReadModbus := FALSE; END_IF;
   #_w1 := #PH_xEndWriteModbus;
   IF #_w1 THEN
       #PH_xEndWriteModbus := FALSE;
       #PH_xReadModbus := TRUE;
   END_IF;
END_REGION

REGION Network 33 (SCL): ### HMI STATUS ###
   IF #ST_xStoppingFaults THEN
       #tHMR.dStatus := 7;
   ELSIF #AUX_rgtIN_tDriveData.rgxStatusBits.xStatus_MoveProgress OR (#IN_xSimulationActive AND #AUX_dSimWaitEnd_ms > 0) THEN
       #tHMR.dStatus := 3;
   ELSE
       #tHMR.dStatus := 1;
   END_IF;

   IF #tHMR.dXCutStatusRequest = 3 AND #AUX_rgtIN_tDriveData.rgxStatusBits.xStatus_BridgeEnabled THEN
       #tHMR.dXCutActualStatus := 3;
   ELSE
       #tHMR.dXCutActualStatus := 1;

   END_IF;

   IF NOT #IN_xSimulationActive THEN
       #tHMR.dCarriagePosition_cmm := #AUX_rgtIN_tDriveData.dCarriagePos_dmm * 10;
   END_IF;

   #tHMR.dTimeHeadDown_ms := INT_TO_DINT(#AUX_rgtIN_tDriveData.iTimeHeadDown_ms);
END_REGION

REGION Network 34: ####_OUTPUT_####
END_REGION

REGION Network 35: Enable / disable bridge
   RUNG wire#powerrail
      { S7_Templates := "SrcType := DInt" } EQ_Contact(in1 := #tHMR.dXCutStatusRequest, in2 := #CONST_DENABLED)
      Coil( #AUX_tOutputDrive.rgxControlBits.xEnableBridge )
   END_RUNG
   RUNG wire#powerrail
      { S7_Templates := "SrcType := DInt" } EQ_Contact(in1 := #tHMR.dXCutStatusRequest, in2 := #CONST_DDISABLED)
      Coil( #AUX_tOutputDrive.rgxControlBits.xDisableBridge )
   END_RUNG
   // the same network as SCL:
   #AUX_tOutputDrive.rgxControlBits.xEnableBridge := #tHMR.dXCutStatusRequest = #CONST_DENABLED;
   #AUX_tOutputDrive.rgxControlBits.xDisableBridge := #tHMR.dXCutStatusRequest = #CONST_DDISABLED;
END_REGION

REGION Network 36: Simulation mode
   RUNG wire#powerrail
      Contact( FALSE )
      Coil( #AUX_tOutputDrive.rgxControlBits.xSimulationMode )
   END_RUNG
   // the same network as SCL:
   #AUX_tOutputDrive.rgxControlBits.xSimulationMode := FALSE;
END_REGION

REGION Network 37: Fault reset
   RUNG wire#powerrail
      Contact( #IN_xResetAlarms )
      Coil( #AUX_tOutputDrive.rgxControlBits.xFaultReset )
   END_RUNG
   // the same network as SCL:
   #AUX_tOutputDrive.rgxControlBits.xFaultReset := #IN_xResetAlarms;
END_REGION

REGION Network 38 (SCL): Update data to inverter
   #AUX_rgtOUT_tDriveData.dBridgeAngle_degre_10000 := #tHMR.dAngleValue_uDegree / 100;

   IF #AUX_dCutStartPosUp_cmm < #AUX_dCutStartPosDw_cmm THEN
       #AUX_rgtOUT_tDriveData.dHeadDownPos_dmm := #AUX_dCutStartPosUp_cmm / 10;
   ELSE
       #AUX_rgtOUT_tDriveData.dHeadDownPos_dmm := #AUX_dCutStartPosDw_cmm / 10;
   END_IF;

   IF #AUX_dCutStopPosUp_cmm > #AUX_dCutStopPosDw_cmm THEN
       #AUX_rgtOUT_tDriveData.dHeadRisePos_dmm := #AUX_dCutStopPosUp_cmm / 10;
   ELSE
       #AUX_rgtOUT_tDriveData.dHeadRisePos_dmm := #AUX_dCutStopPosDw_cmm / 10;
   END_IF;

   IF #AUX_dNextPlateTime_ms > #AUX_dCutTime20Per_ms THEN
       #AUX_rgtOUT_tDriveData.iReturnSpeed_rpm := REAL_TO_INT(DINT_TO_REAL(#CONST_DMAXRETSPEED_RPM) * 0.2);
   ELSIF #AUX_dNextPlateTime_ms > #AUX_dCutTime40Per_ms THEN
       #AUX_rgtOUT_tDriveData.iReturnSpeed_rpm := REAL_TO_INT(DINT_TO_REAL(#CONST_DMAXRETSPEED_RPM) * 0.4);
   ELSIF #AUX_dNextPlateTime_ms > #AUX_dCutTime60Per_ms THEN
       #AUX_rgtOUT_tDriveData.iReturnSpeed_rpm := REAL_TO_INT(DINT_TO_REAL(#CONST_DMAXRETSPEED_RPM) * 0.6);
   ELSIF #AUX_dNextPlateTime_ms > #AUX_dCutTime80Per_ms THEN
       #AUX_rgtOUT_tDriveData.iReturnSpeed_rpm := REAL_TO_INT(DINT_TO_REAL(#CONST_DMAXRETSPEED_RPM) * 0.8);
   ELSIF #AUX_dNextPlateTime_ms > #AUX_dCutTime100Per_ms THEN
       #AUX_rgtOUT_tDriveData.iReturnSpeed_rpm := REAL_TO_INT(#CONST_DMAXRETSPEED_RPM);
   ELSE
       #AUX_rgtOUT_tDriveData.iReturnSpeed_rpm := 3750;
   END_IF;

   #AUX_rgtOUT_tDriveData.iTimeHeadDown_ms := DINT_TO_INT(#tHMW.dDescReactTime_ms);
   #AUX_rgtOUT_tDriveData.iTimeHeadUp_ms := DINT_TO_INT(#tHMW.dRaiseReactTime_ms);
   #AUX_rgtOUT_tDriveData.iLubAdvanceTime_ms := DINT_TO_INT(#tHMW.dOilONDelay_ms * -1);
   #AUX_rgtOUT_tDriveData.iLubDelayTime_ms := DINT_TO_INT(#tHMW.dOilOFFDelay_ms);
   #AUX_rgtOUT_tDriveData.iTimeHeadAct_ms := DINT_TO_INT(#tHMW.dFireONReactTime_ms);
   #AUX_rgtOUT_tDriveData.iTimeHeadDeactiv_ms := DINT_TO_INT(#tHMW.dFireOFFReactTime_ms);
   #AUX_rgtOUT_tDriveData.dPressure_mN := #tHMW.dCuttingPressure_mN;
   #AUX_rgtOUT_tDriveData.dMissionID := #AUX_dMissionToSend;
   #AUX_rgtOUT_tDriveData.dMissionCounter := #AUX_dMissionCounterValue_cmm;

   IF #INO_tEnc.rgxMetersForXcuts[#IN_dXCutIndex] THEN

       #AUX_rgtOUT_tDriveData.dSyncroCounter := #INO_tEnc.dLastMeterValue_cmm;
       #INO_tEnc.rgxMetersForXcuts[#IN_dXCutIndex] := FALSE;

   END_IF;